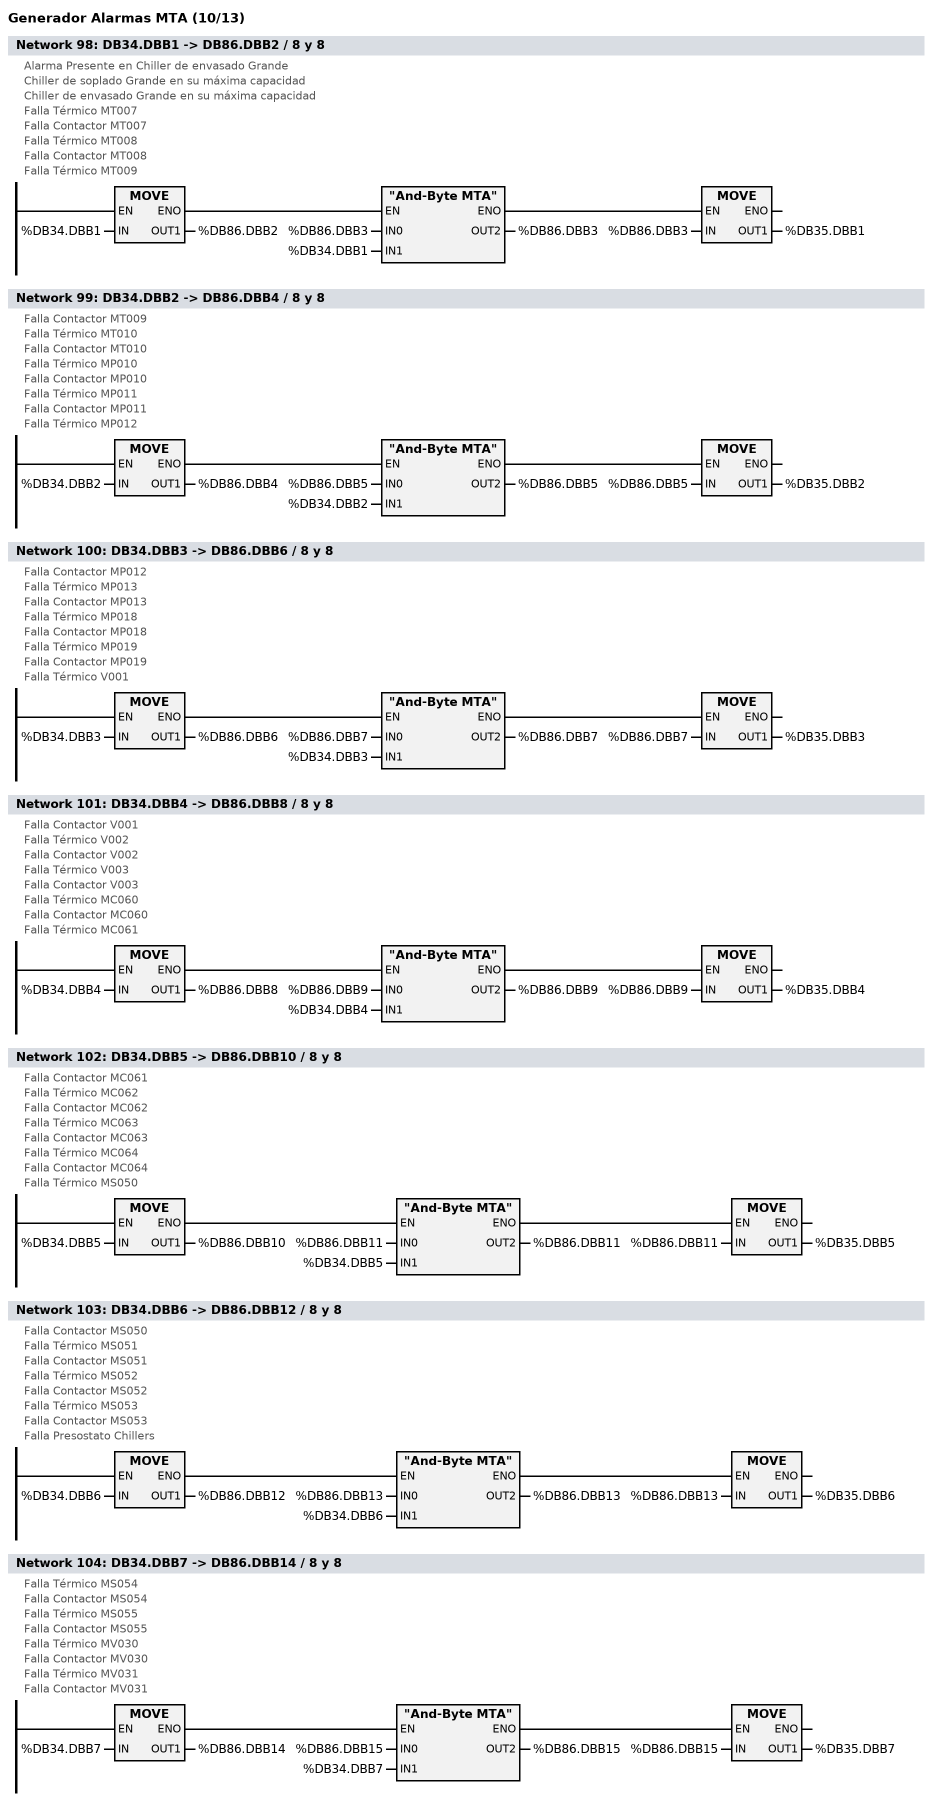
   RUNG wire#powerrail
      { S7_GenerateENO := "TRUE" } Move(in := %DB34.DBB1, out1 => %DB86.DBB2)
      "And-Byte MTA"(IN0 := %DB86.DBB3, IN1 := %DB34.DBB1, OUT2 => %DB86.DBB3)
      { S7_GenerateENO := "TRUE" } Move(in := %DB86.DBB3, out1 => %DB35.DBB1)
   END_RUNG
   // the same network as SCL:
   // ENO of a box is taken as its EN; it also drops when the box reports an error
   %DB86.DBB2 := %DB34.DBB1;
   "And-Byte MTA"(IN0 := %DB86.DBB3, IN1 := %DB34.DBB1, OUT2 => %DB86.DBB3, ENO => #_w1);
   IF #_w1 THEN %DB35.DBB1 := %DB86.DBB3; END_IF;
END_REGION

REGION Network 99: DB34.DBB2 -> DB86.DBB4 / 8 y 8
   // Falla Contactor MT009
   // Falla Térmico MT010
   // Falla Contactor MT010
   // Falla Térmico MP010
   // Falla Contactor MP010
   // Falla Térmico MP011
   // Falla Contactor MP011
   // Falla Térmico MP012
   RUNG wire#powerrail
      { S7_GenerateENO := "TRUE" } Move(in := %DB34.DBB2, out1 => %DB86.DBB4)
      "And-Byte MTA"(IN0 := %DB86.DBB5, IN1 := %DB34.DBB2, OUT2 => %DB86.DBB5)
      { S7_GenerateENO := "TRUE" } Move(in := %DB86.DBB5, out1 => %DB35.DBB2)
   END_RUNG
   // the same network as SCL:
   // ENO of a box is taken as its EN; it also drops when the box reports an error
   %DB86.DBB4 := %DB34.DBB2;
   "And-Byte MTA"(IN0 := %DB86.DBB5, IN1 := %DB34.DBB2, OUT2 => %DB86.DBB5, ENO => #_w1);
   IF #_w1 THEN %DB35.DBB2 := %DB86.DBB5; END_IF;
END_REGION

REGION Network 100: DB34.DBB3 -> DB86.DBB6 / 8 y 8
   // Falla Contactor MP012
   // Falla Térmico MP013
   // Falla Contactor MP013
   // Falla Térmico MP018
   // Falla Contactor MP018
   // Falla Térmico MP019
   // Falla Contactor MP019
   // Falla Térmico V001
   RUNG wire#powerrail
      { S7_GenerateENO := "TRUE" } Move(in := %DB34.DBB3, out1 => %DB86.DBB6)
      "And-Byte MTA"(IN0 := %DB86.DBB7, IN1 := %DB34.DBB3, OUT2 => %DB86.DBB7)
      { S7_GenerateENO := "TRUE" } Move(in := %DB86.DBB7, out1 => %DB35.DBB3)
   END_RUNG
   // the same network as SCL:
   // ENO of a box is taken as its EN; it also drops when the box reports an error
   %DB86.DBB6 := %DB34.DBB3;
   "And-Byte MTA"(IN0 := %DB86.DBB7, IN1 := %DB34.DBB3, OUT2 => %DB86.DBB7, ENO => #_w1);
   IF #_w1 THEN %DB35.DBB3 := %DB86.DBB7; END_IF;
END_REGION

REGION Network 101: DB34.DBB4 -> DB86.DBB8 / 8 y 8
   // Falla Contactor V001
   // Falla Térmico V002
   // Falla Contactor V002
   // Falla Térmico V003
   // Falla Contactor V003
   // Falla Térmico MC060
   // Falla Contactor MC060
   // Falla Térmico MC061
   RUNG wire#powerrail
      { S7_GenerateENO := "TRUE" } Move(in := %DB34.DBB4, out1 => %DB86.DBB8)
      "And-Byte MTA"(IN0 := %DB86.DBB9, IN1 := %DB34.DBB4, OUT2 => %DB86.DBB9)
      { S7_GenerateENO := "TRUE" } Move(in := %DB86.DBB9, out1 => %DB35.DBB4)
   END_RUNG
   // the same network as SCL:
   // ENO of a box is taken as its EN; it also drops when the box reports an error
   %DB86.DBB8 := %DB34.DBB4;
   "And-Byte MTA"(IN0 := %DB86.DBB9, IN1 := %DB34.DBB4, OUT2 => %DB86.DBB9, ENO => #_w1);
   IF #_w1 THEN %DB35.DBB4 := %DB86.DBB9; END_IF;
END_REGION

REGION Network 102: DB34.DBB5 -> DB86.DBB10 / 8 y 8
   // Falla Contactor MC061
   // Falla Térmico MC062
   // Falla Contactor MC062
   // Falla Térmico MC063
   // Falla Contactor MC063
   // Falla Térmico MC064
   // Falla Contactor MC064
   // Falla Térmico MS050
   RUNG wire#powerrail
      { S7_GenerateENO := "TRUE" } Move(in := %DB34.DBB5, out1 => %DB86.DBB10)
      "And-Byte MTA"(IN0 := %DB86.DBB11, IN1 := %DB34.DBB5, OUT2 => %DB86.DBB11)
      { S7_GenerateENO := "TRUE" } Move(in := %DB86.DBB11, out1 => %DB35.DBB5)
   END_RUNG
   // the same network as SCL:
   // ENO of a box is taken as its EN; it also drops when the box reports an error
   %DB86.DBB10 := %DB34.DBB5;
   "And-Byte MTA"(IN0 := %DB86.DBB11, IN1 := %DB34.DBB5, OUT2 => %DB86.DBB11, ENO => #_w1);
   IF #_w1 THEN %DB35.DBB5 := %DB86.DBB11; END_IF;
END_REGION

REGION Network 103: DB34.DBB6 -> DB86.DBB12 / 8 y 8
   // Falla Contactor MS050
   // Falla Térmico MS051
   // Falla Contactor MS051
   // Falla Térmico MS052
   // Falla Contactor MS052
   // Falla Térmico MS053
   // Falla Contactor MS053
   // Falla Presostato Chillers
   RUNG wire#powerrail
      { S7_GenerateENO := "TRUE" } Move(in := %DB34.DBB6, out1 => %DB86.DBB12)
      "And-Byte MTA"(IN0 := %DB86.DBB13, IN1 := %DB34.DBB6, OUT2 => %DB86.DBB13)
      { S7_GenerateENO := "TRUE" } Move(in := %DB86.DBB13, out1 => %DB35.DBB6)
   END_RUNG
   // the same network as SCL:
   // ENO of a box is taken as its EN; it also drops when the box reports an error
   %DB86.DBB12 := %DB34.DBB6;
   "And-Byte MTA"(IN0 := %DB86.DBB13, IN1 := %DB34.DBB6, OUT2 => %DB86.DBB13, ENO => #_w1);
   IF #_w1 THEN %DB35.DBB6 := %DB86.DBB13; END_IF;
END_REGION

REGION Network 104: DB34.DBB7 -> DB86.DBB14 / 8 y 8
   // Falla Térmico MS054
   // Falla Contactor MS054
   // Falla Térmico MS055
   // Falla Contactor MS055
   // Falla Térmico MV030
   // Falla Contactor MV030
   // Falla Térmico MV031
   // Falla Contactor MV031
   RUNG wire#powerrail
      { S7_GenerateENO := "TRUE" } Move(in := %DB34.DBB7, out1 => %DB86.DBB14)
      "And-Byte MTA"(IN0 := %DB86.DBB15, IN1 := %DB34.DBB7, OUT2 => %DB86.DBB15)
      { S7_GenerateENO := "TRUE" } Move(in := %DB86.DBB15, out1 => %DB35.DBB7)
   END_RUNG
   // the same network as SCL:
   // ENO of a box is taken as its EN; it also drops when the box reports an error
   %DB86.DBB14 := %DB34.DBB7;
   "And-Byte MTA"(IN0 := %DB86.DBB15, IN1 := %DB34.DBB7, OUT2 => %DB86.DBB15, ENO => #_w1);
   IF #_w1 THEN %DB35.DBB7 := %DB86.DBB15; END_IF;
END_REGION

REGION Network 105: DB34.DBB8 -> DB86.DBB16 / 8 y 8
   // Falla Térmico MP014
   // Falla Contactor MP014
   // Falla Térmico MP015
   // Falla Contactor MP015
   // Falla Térmico MC001
   // Falla Contactor MC001
   // Falla Térmico MC002
   // Falla Contactor MC002
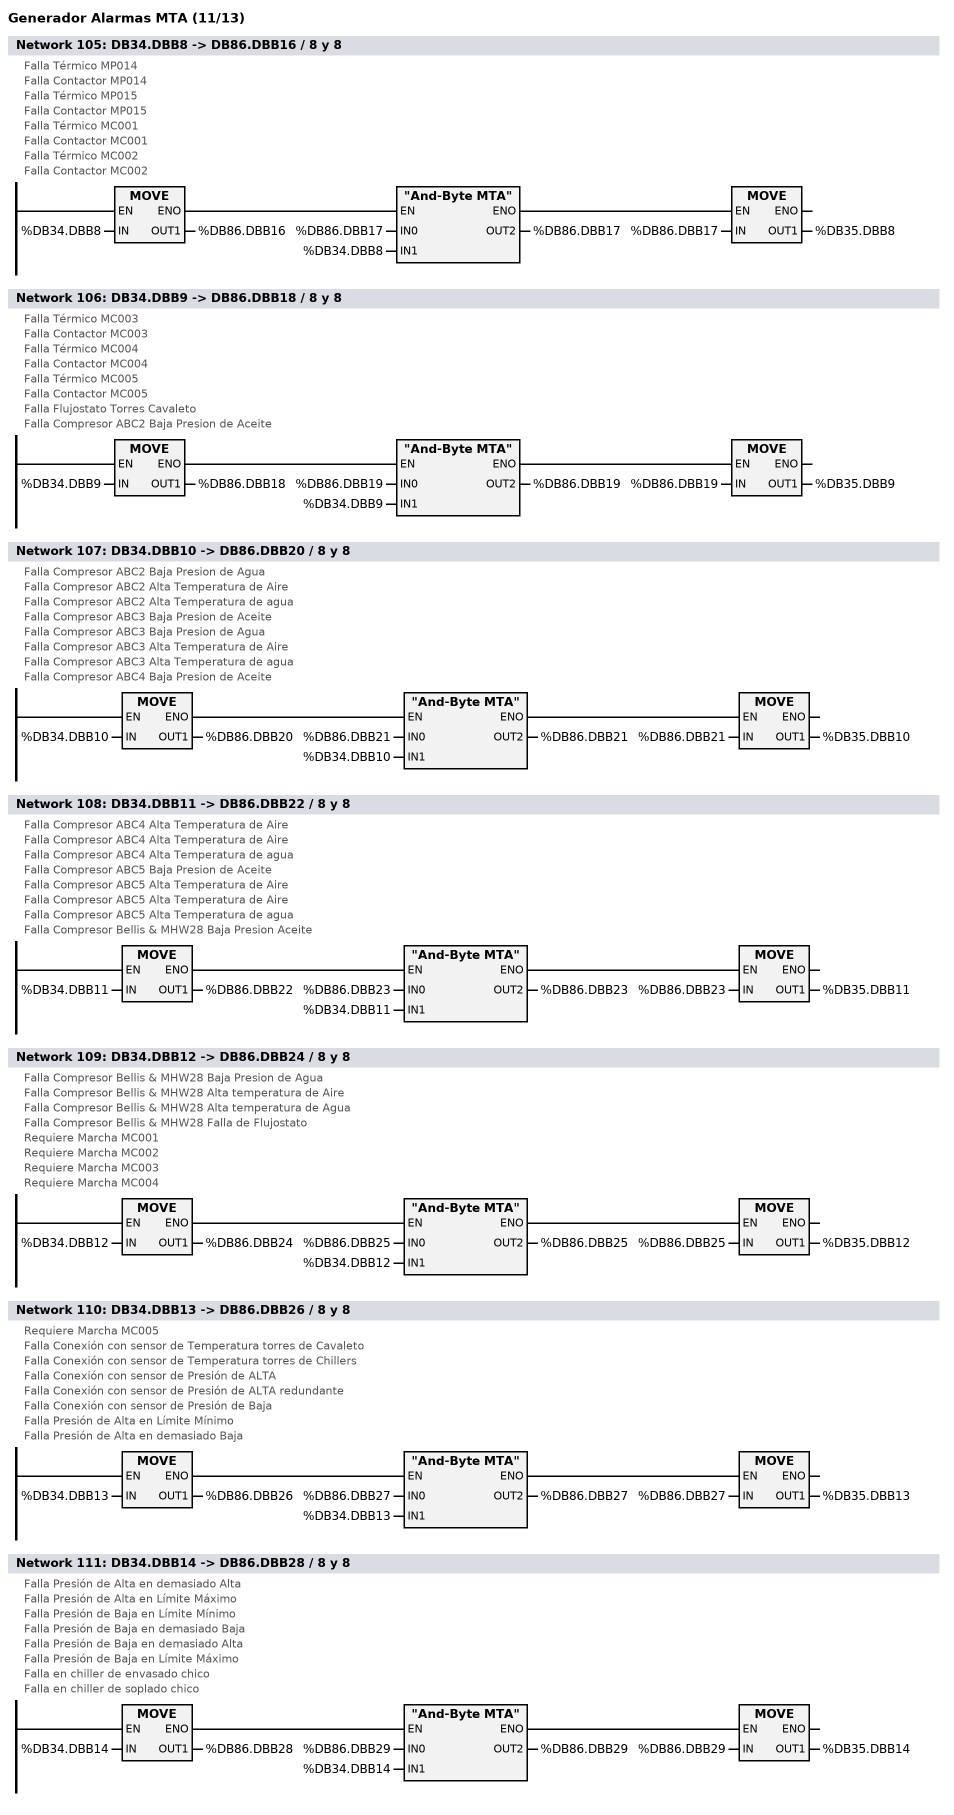
   RUNG wire#powerrail
      { S7_GenerateENO := "TRUE" } Move(in := %DB34.DBB8, out1 => %DB86.DBB16)
      "And-Byte MTA"(IN0 := %DB86.DBB17, IN1 := %DB34.DBB8, OUT2 => %DB86.DBB17)
      { S7_GenerateENO := "TRUE" } Move(in := %DB86.DBB17, out1 => %DB35.DBB8)
   END_RUNG
   // the same network as SCL:
   // ENO of a box is taken as its EN; it also drops when the box reports an error
   %DB86.DBB16 := %DB34.DBB8;
   "And-Byte MTA"(IN0 := %DB86.DBB17, IN1 := %DB34.DBB8, OUT2 => %DB86.DBB17, ENO => #_w1);
   IF #_w1 THEN %DB35.DBB8 := %DB86.DBB17; END_IF;
END_REGION

REGION Network 106: DB34.DBB9 -> DB86.DBB18 / 8 y 8
   // Falla Térmico MC003
   // Falla Contactor MC003
   // Falla Térmico MC004
   // Falla Contactor MC004
   // Falla Térmico MC005
   // Falla Contactor MC005
   // Falla Flujostato Torres Cavaleto
   // Falla Compresor ABC2 Baja Presion de Aceite
   RUNG wire#powerrail
      { S7_GenerateENO := "TRUE" } Move(in := %DB34.DBB9, out1 => %DB86.DBB18)
      "And-Byte MTA"(IN0 := %DB86.DBB19, IN1 := %DB34.DBB9, OUT2 => %DB86.DBB19)
      { S7_GenerateENO := "TRUE" } Move(in := %DB86.DBB19, out1 => %DB35.DBB9)
   END_RUNG
   // the same network as SCL:
   // ENO of a box is taken as its EN; it also drops when the box reports an error
   %DB86.DBB18 := %DB34.DBB9;
   "And-Byte MTA"(IN0 := %DB86.DBB19, IN1 := %DB34.DBB9, OUT2 => %DB86.DBB19, ENO => #_w1);
   IF #_w1 THEN %DB35.DBB9 := %DB86.DBB19; END_IF;
END_REGION

REGION Network 107: DB34.DBB10 -> DB86.DBB20 / 8 y 8
   // Falla Compresor ABC2 Baja Presion de Agua
   // Falla Compresor ABC2 Alta Temperatura de Aire
   // Falla Compresor ABC2 Alta Temperatura de agua
   // Falla Compresor ABC3 Baja Presion de Aceite
   // Falla Compresor ABC3 Baja Presion de Agua
   // Falla Compresor ABC3 Alta Temperatura de Aire
   // Falla Compresor ABC3 Alta Temperatura de agua
   // Falla Compresor ABC4 Baja Presion de Aceite
   RUNG wire#powerrail
      { S7_GenerateENO := "TRUE" } Move(in := %DB34.DBB10, out1 => %DB86.DBB20)
      "And-Byte MTA"(IN0 := %DB86.DBB21, IN1 := %DB34.DBB10, OUT2 => %DB86.DBB21)
      { S7_GenerateENO := "TRUE" } Move(in := %DB86.DBB21, out1 => %DB35.DBB10)
   END_RUNG
   // the same network as SCL:
   // ENO of a box is taken as its EN; it also drops when the box reports an error
   %DB86.DBB20 := %DB34.DBB10;
   "And-Byte MTA"(IN0 := %DB86.DBB21, IN1 := %DB34.DBB10, OUT2 => %DB86.DBB21, ENO => #_w1);
   IF #_w1 THEN %DB35.DBB10 := %DB86.DBB21; END_IF;
END_REGION

REGION Network 108: DB34.DBB11 -> DB86.DBB22 / 8 y 8
   // Falla Compresor ABC4 Alta Temperatura de Aire
   // Falla Compresor ABC4 Alta Temperatura de Aire
   // Falla Compresor ABC4 Alta Temperatura de agua
   // Falla Compresor ABC5 Baja Presion de Aceite
   // Falla Compresor ABC5 Alta Temperatura de Aire
   // Falla Compresor ABC5 Alta Temperatura de Aire
   // Falla Compresor ABC5 Alta Temperatura de agua
   // Falla Compresor Bellis & MHW28 Baja Presion Aceite
   RUNG wire#powerrail
      { S7_GenerateENO := "TRUE" } Move(in := %DB34.DBB11, out1 => %DB86.DBB22)
      "And-Byte MTA"(IN0 := %DB86.DBB23, IN1 := %DB34.DBB11, OUT2 => %DB86.DBB23)
      { S7_GenerateENO := "TRUE" } Move(in := %DB86.DBB23, out1 => %DB35.DBB11)
   END_RUNG
   // the same network as SCL:
   // ENO of a box is taken as its EN; it also drops when the box reports an error
   %DB86.DBB22 := %DB34.DBB11;
   "And-Byte MTA"(IN0 := %DB86.DBB23, IN1 := %DB34.DBB11, OUT2 => %DB86.DBB23, ENO => #_w1);
   IF #_w1 THEN %DB35.DBB11 := %DB86.DBB23; END_IF;
END_REGION

REGION Network 109: DB34.DBB12 -> DB86.DBB24 / 8 y 8
   // Falla Compresor Bellis & MHW28 Baja Presion de Agua
   // Falla Compresor Bellis & MHW28 Alta temperatura de Aire
   // Falla Compresor Bellis & MHW28 Alta temperatura de Agua
   // Falla Compresor Bellis & MHW28 Falla de Flujostato
   // Requiere Marcha MC001
   // Requiere Marcha MC002
   // Requiere Marcha MC003
   // Requiere Marcha MC004
   RUNG wire#powerrail
      { S7_GenerateENO := "TRUE" } Move(in := %DB34.DBB12, out1 => %DB86.DBB24)
      "And-Byte MTA"(IN0 := %DB86.DBB25, IN1 := %DB34.DBB12, OUT2 => %DB86.DBB25)
      { S7_GenerateENO := "TRUE" } Move(in := %DB86.DBB25, out1 => %DB35.DBB12)
   END_RUNG
   // the same network as SCL:
   // ENO of a box is taken as its EN; it also drops when the box reports an error
   %DB86.DBB24 := %DB34.DBB12;
   "And-Byte MTA"(IN0 := %DB86.DBB25, IN1 := %DB34.DBB12, OUT2 => %DB86.DBB25, ENO => #_w1);
   IF #_w1 THEN %DB35.DBB12 := %DB86.DBB25; END_IF;
END_REGION

REGION Network 110: DB34.DBB13 -> DB86.DBB26 / 8 y 8
   // Requiere Marcha MC005
   // Falla Conexión con sensor de Temperatura torres de Cavaleto
   // Falla Conexión con sensor de Temperatura torres de Chillers
   // Falla Conexión con sensor de Presión de ALTA
   // Falla Conexión con sensor de Presión de ALTA redundante
   // Falla Conexión con sensor de Presión de Baja
   // Falla Presión de Alta en Límite Mínimo
   // Falla Presión de Alta en demasiado Baja
   RUNG wire#powerrail
      { S7_GenerateENO := "TRUE" } Move(in := %DB34.DBB13, out1 => %DB86.DBB26)
      "And-Byte MTA"(IN0 := %DB86.DBB27, IN1 := %DB34.DBB13, OUT2 => %DB86.DBB27)
      { S7_GenerateENO := "TRUE" } Move(in := %DB86.DBB27, out1 => %DB35.DBB13)
   END_RUNG
   // the same network as SCL:
   // ENO of a box is taken as its EN; it also drops when the box reports an error
   %DB86.DBB26 := %DB34.DBB13;
   "And-Byte MTA"(IN0 := %DB86.DBB27, IN1 := %DB34.DBB13, OUT2 => %DB86.DBB27, ENO => #_w1);
   IF #_w1 THEN %DB35.DBB13 := %DB86.DBB27; END_IF;
END_REGION

REGION Network 111: DB34.DBB14 -> DB86.DBB28 / 8 y 8
   // Falla Presión de Alta en demasiado Alta
   // Falla Presión de Alta en Límite Máximo
   // Falla Presión de Baja en Límite Mínimo
   // Falla Presión de Baja en demasiado Baja
   // Falla Presión de Baja en demasiado Alta
   // Falla Presión de Baja en Límite Máximo
   // Falla en chiller de envasado chico
   // Falla en chiller de soplado chico
   RUNG wire#powerrail
      { S7_GenerateENO := "TRUE" } Move(in := %DB34.DBB14, out1 => %DB86.DBB28)
      "And-Byte MTA"(IN0 := %DB86.DBB29, IN1 := %DB34.DBB14, OUT2 => %DB86.DBB29)
      { S7_GenerateENO := "TRUE" } Move(in := %DB86.DBB29, out1 => %DB35.DBB14)
   END_RUNG
   // the same network as SCL:
   // ENO of a box is taken as its EN; it also drops when the box reports an error
   %DB86.DBB28 := %DB34.DBB14;
   "And-Byte MTA"(IN0 := %DB86.DBB29, IN1 := %DB34.DBB14, OUT2 => %DB86.DBB29, ENO => #_w1);
   IF #_w1 THEN %DB35.DBB14 := %DB86.DBB29; END_IF;
END_REGION

REGION Network 112: DB34.DBB15 -> DB86.DBB30 / 8 y 8
   // Horas máximas en Compresor 1
   // Horas máximas en Compresor 2
   // Horas máximas en Compresor 3
   // Horas máximas en Compresor 4
   // Horas máximas en Compresor 5
   // Falla algún contactor en Booster 1
   // Falla algún guardamotor en Booster 1
   // Presión Alta en Booster
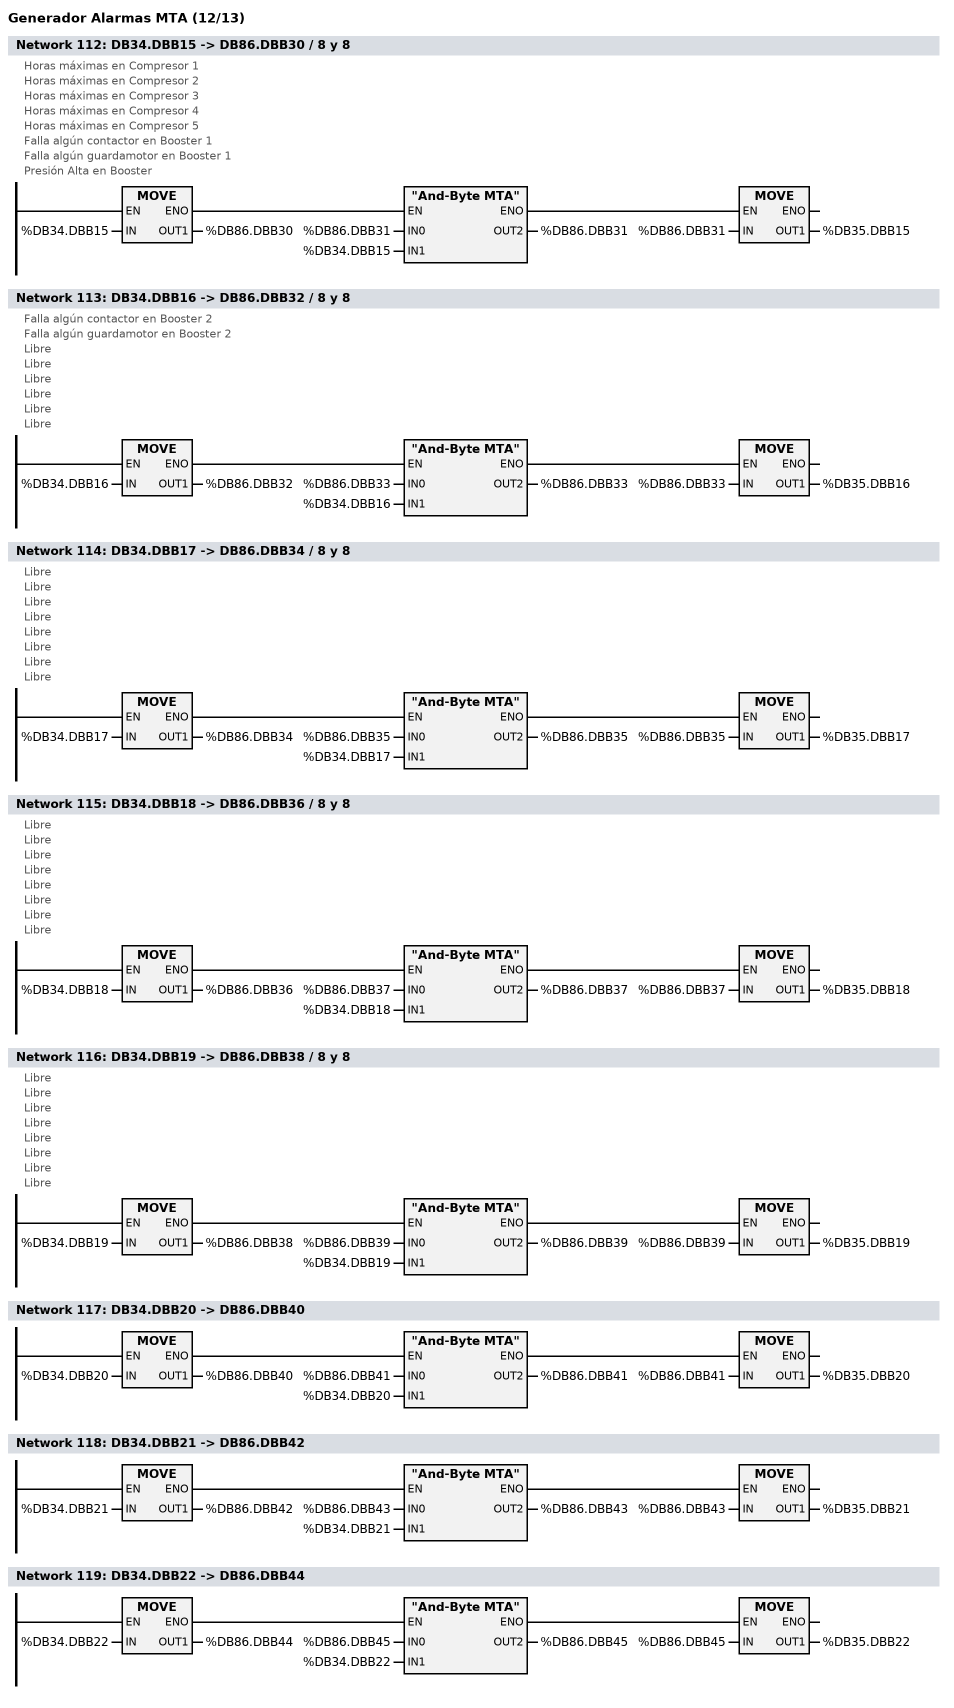
   RUNG wire#powerrail
      { S7_GenerateENO := "TRUE" } Move(in := %DB34.DBB15, out1 => %DB86.DBB30)
      "And-Byte MTA"(IN0 := %DB86.DBB31, IN1 := %DB34.DBB15, OUT2 => %DB86.DBB31)
      { S7_GenerateENO := "TRUE" } Move(in := %DB86.DBB31, out1 => %DB35.DBB15)
   END_RUNG
   // the same network as SCL:
   // ENO of a box is taken as its EN; it also drops when the box reports an error
   %DB86.DBB30 := %DB34.DBB15;
   "And-Byte MTA"(IN0 := %DB86.DBB31, IN1 := %DB34.DBB15, OUT2 => %DB86.DBB31, ENO => #_w1);
   IF #_w1 THEN %DB35.DBB15 := %DB86.DBB31; END_IF;
END_REGION

REGION Network 113: DB34.DBB16 -> DB86.DBB32 / 8 y 8
   // Falla algún contactor en Booster 2
   // Falla algún guardamotor en Booster 2
   // Libre
   // Libre
   // Libre
   // Libre
   // Libre
   // Libre
   RUNG wire#powerrail
      { S7_GenerateENO := "TRUE" } Move(in := %DB34.DBB16, out1 => %DB86.DBB32)
      "And-Byte MTA"(IN0 := %DB86.DBB33, IN1 := %DB34.DBB16, OUT2 => %DB86.DBB33)
      { S7_GenerateENO := "TRUE" } Move(in := %DB86.DBB33, out1 => %DB35.DBB16)
   END_RUNG
   // the same network as SCL:
   // ENO of a box is taken as its EN; it also drops when the box reports an error
   %DB86.DBB32 := %DB34.DBB16;
   "And-Byte MTA"(IN0 := %DB86.DBB33, IN1 := %DB34.DBB16, OUT2 => %DB86.DBB33, ENO => #_w1);
   IF #_w1 THEN %DB35.DBB16 := %DB86.DBB33; END_IF;
END_REGION

REGION Network 114: DB34.DBB17 -> DB86.DBB34 / 8 y 8
   // Libre
   // Libre
   // Libre
   // Libre
   // Libre
   // Libre
   // Libre
   // Libre
   RUNG wire#powerrail
      { S7_GenerateENO := "TRUE" } Move(in := %DB34.DBB17, out1 => %DB86.DBB34)
      "And-Byte MTA"(IN0 := %DB86.DBB35, IN1 := %DB34.DBB17, OUT2 => %DB86.DBB35)
      { S7_GenerateENO := "TRUE" } Move(in := %DB86.DBB35, out1 => %DB35.DBB17)
   END_RUNG
   // the same network as SCL:
   // ENO of a box is taken as its EN; it also drops when the box reports an error
   %DB86.DBB34 := %DB34.DBB17;
   "And-Byte MTA"(IN0 := %DB86.DBB35, IN1 := %DB34.DBB17, OUT2 => %DB86.DBB35, ENO => #_w1);
   IF #_w1 THEN %DB35.DBB17 := %DB86.DBB35; END_IF;
END_REGION

REGION Network 115: DB34.DBB18 -> DB86.DBB36 / 8 y 8
   // Libre
   // Libre
   // Libre
   // Libre
   // Libre
   // Libre
   // Libre
   // Libre
   RUNG wire#powerrail
      { S7_GenerateENO := "TRUE" } Move(in := %DB34.DBB18, out1 => %DB86.DBB36)
      "And-Byte MTA"(IN0 := %DB86.DBB37, IN1 := %DB34.DBB18, OUT2 => %DB86.DBB37)
      { S7_GenerateENO := "TRUE" } Move(in := %DB86.DBB37, out1 => %DB35.DBB18)
   END_RUNG
   // the same network as SCL:
   // ENO of a box is taken as its EN; it also drops when the box reports an error
   %DB86.DBB36 := %DB34.DBB18;
   "And-Byte MTA"(IN0 := %DB86.DBB37, IN1 := %DB34.DBB18, OUT2 => %DB86.DBB37, ENO => #_w1);
   IF #_w1 THEN %DB35.DBB18 := %DB86.DBB37; END_IF;
END_REGION

REGION Network 116: DB34.DBB19 -> DB86.DBB38 / 8 y 8
   // Libre
   // Libre
   // Libre
   // Libre
   // Libre
   // Libre
   // Libre
   // Libre
   RUNG wire#powerrail
      { S7_GenerateENO := "TRUE" } Move(in := %DB34.DBB19, out1 => %DB86.DBB38)
      "And-Byte MTA"(IN0 := %DB86.DBB39, IN1 := %DB34.DBB19, OUT2 => %DB86.DBB39)
      { S7_GenerateENO := "TRUE" } Move(in := %DB86.DBB39, out1 => %DB35.DBB19)
   END_RUNG
   // the same network as SCL:
   // ENO of a box is taken as its EN; it also drops when the box reports an error
   %DB86.DBB38 := %DB34.DBB19;
   "And-Byte MTA"(IN0 := %DB86.DBB39, IN1 := %DB34.DBB19, OUT2 => %DB86.DBB39, ENO => #_w1);
   IF #_w1 THEN %DB35.DBB19 := %DB86.DBB39; END_IF;
END_REGION

REGION Network 117: DB34.DBB20 -> DB86.DBB40
   RUNG wire#powerrail
      { S7_GenerateENO := "TRUE" } Move(in := %DB34.DBB20, out1 => %DB86.DBB40)
      "And-Byte MTA"(IN0 := %DB86.DBB41, IN1 := %DB34.DBB20, OUT2 => %DB86.DBB41)
      { S7_GenerateENO := "TRUE" } Move(in := %DB86.DBB41, out1 => %DB35.DBB20)
   END_RUNG
   // the same network as SCL:
   // ENO of a box is taken as its EN; it also drops when the box reports an error
   %DB86.DBB40 := %DB34.DBB20;
   "And-Byte MTA"(IN0 := %DB86.DBB41, IN1 := %DB34.DBB20, OUT2 => %DB86.DBB41, ENO => #_w1);
   IF #_w1 THEN %DB35.DBB20 := %DB86.DBB41; END_IF;
END_REGION

REGION Network 118: DB34.DBB21 -> DB86.DBB42
   RUNG wire#powerrail
      { S7_GenerateENO := "TRUE" } Move(in := %DB34.DBB21, out1 => %DB86.DBB42)
      "And-Byte MTA"(IN0 := %DB86.DBB43, IN1 := %DB34.DBB21, OUT2 => %DB86.DBB43)
      { S7_GenerateENO := "TRUE" } Move(in := %DB86.DBB43, out1 => %DB35.DBB21)
   END_RUNG
   // the same network as SCL:
   // ENO of a box is taken as its EN; it also drops when the box reports an error
   %DB86.DBB42 := %DB34.DBB21;
   "And-Byte MTA"(IN0 := %DB86.DBB43, IN1 := %DB34.DBB21, OUT2 => %DB86.DBB43, ENO => #_w1);
   IF #_w1 THEN %DB35.DBB21 := %DB86.DBB43; END_IF;
END_REGION

REGION Network 119: DB34.DBB22 -> DB86.DBB44
   RUNG wire#powerrail
      { S7_GenerateENO := "TRUE" } Move(in := %DB34.DBB22, out1 => %DB86.DBB44)
      "And-Byte MTA"(IN0 := %DB86.DBB45, IN1 := %DB34.DBB22, OUT2 => %DB86.DBB45)
      { S7_GenerateENO := "TRUE" } Move(in := %DB86.DBB45, out1 => %DB35.DBB22)
   END_RUNG
   // the same network as SCL:
   // ENO of a box is taken as its EN; it also drops when the box reports an error
   %DB86.DBB44 := %DB34.DBB22;
   "And-Byte MTA"(IN0 := %DB86.DBB45, IN1 := %DB34.DBB22, OUT2 => %DB86.DBB45, ENO => #_w1);
   IF #_w1 THEN %DB35.DBB22 := %DB86.DBB45; END_IF;
END_REGION

REGION Network 120: DB34.DBB23 -> DB86.DBB46
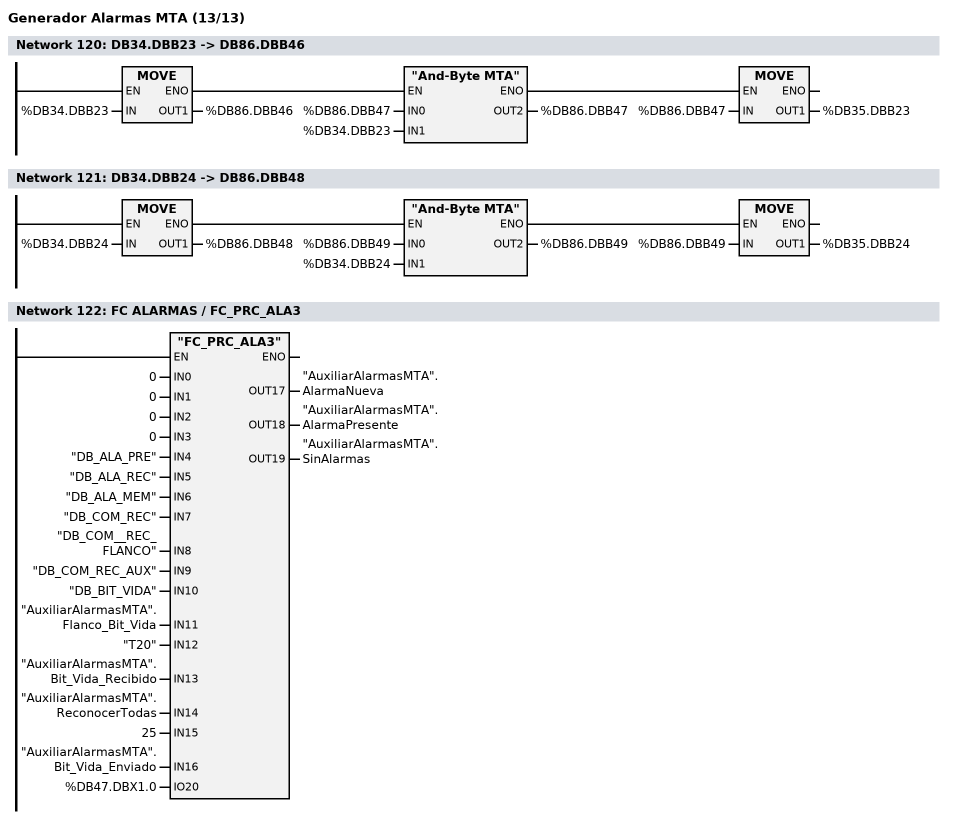
   RUNG wire#powerrail
      { S7_GenerateENO := "TRUE" } Move(in := %DB34.DBB23, out1 => %DB86.DBB46)
      "And-Byte MTA"(IN0 := %DB86.DBB47, IN1 := %DB34.DBB23, OUT2 => %DB86.DBB47)
      { S7_GenerateENO := "TRUE" } Move(in := %DB86.DBB47, out1 => %DB35.DBB23)
   END_RUNG
   // the same network as SCL:
   // ENO of a box is taken as its EN; it also drops when the box reports an error
   %DB86.DBB46 := %DB34.DBB23;
   "And-Byte MTA"(IN0 := %DB86.DBB47, IN1 := %DB34.DBB23, OUT2 => %DB86.DBB47, ENO => #_w1);
   IF #_w1 THEN %DB35.DBB23 := %DB86.DBB47; END_IF;
END_REGION

REGION Network 121: DB34.DBB24 -> DB86.DBB48
   RUNG wire#powerrail
      { S7_GenerateENO := "TRUE" } Move(in := %DB34.DBB24, out1 => %DB86.DBB48)
      "And-Byte MTA"(IN0 := %DB86.DBB49, IN1 := %DB34.DBB24, OUT2 => %DB86.DBB49)
      { S7_GenerateENO := "TRUE" } Move(in := %DB86.DBB49, out1 => %DB35.DBB24)
   END_RUNG
   // the same network as SCL:
   // ENO of a box is taken as its EN; it also drops when the box reports an error
   %DB86.DBB48 := %DB34.DBB24;
   "And-Byte MTA"(IN0 := %DB86.DBB49, IN1 := %DB34.DBB24, OUT2 => %DB86.DBB49, ENO => #_w1);
   IF #_w1 THEN %DB35.DBB24 := %DB86.DBB49; END_IF;
END_REGION

REGION Network 122: FC ALARMAS / FC_PRC_ALA3
   RUNG wire#powerrail
      "FC_PRC_ALA3"(IN0 := 0, IN1 := 0, IN2 := 0, IN3 := 0, IN4 := "DB_ALA_PRE", IN5 := "DB_ALA_REC", IN6 := "DB_ALA_MEM", IN7 := "DB_COM_REC", IN8 := "DB_COM__REC_FLANCO", IN9 := "DB_COM_REC_AUX", IN10 := "DB_BIT_VIDA", IN11 := "AuxiliarAlarmasMTA".Flanco_Bit_Vida, IN12 := "T20", IN13 := "AuxiliarAlarmasMTA".Bit_Vida_Recibido, IN14 := "AuxiliarAlarmasMTA".ReconocerTodas, IN15 := 25, IN16 := "AuxiliarAlarmasMTA".Bit_Vida_Enviado, IO20 := %DB47.DBX1.0, OUT17 => "AuxiliarAlarmasMTA".AlarmaNueva, OUT18 => "AuxiliarAlarmasMTA".AlarmaPresente, OUT19 => "AuxiliarAlarmasMTA".SinAlarmas)
   END_RUNG
   // the same network as SCL:
   "FC_PRC_ALA3"(IN0 := 0,
                 IN1 := 0,
                 IN2 := 0,
                 IN3 := 0,
                 IN4 := "DB_ALA_PRE",
                 IN5 := "DB_ALA_REC",
                 IN6 := "DB_ALA_MEM",
                 IN7 := "DB_COM_REC",
                 IN8 := "DB_COM__REC_FLANCO",
                 IN9 := "DB_COM_REC_AUX",
                 IN10 := "DB_BIT_VIDA",
                 IN11 := "AuxiliarAlarmasMTA".Flanco_Bit_Vida,
                 IN12 := "T20",
                 IN13 := "AuxiliarAlarmasMTA".Bit_Vida_Recibido,
                 IN14 := "AuxiliarAlarmasMTA".ReconocerTodas,
                 IN15 := 25,
                 IN16 := "AuxiliarAlarmasMTA".Bit_Vida_Enviado,
                 IO20 := %DB47.DBX1.0,
                 OUT17 => "AuxiliarAlarmasMTA".AlarmaNueva,
                 OUT18 => "AuxiliarAlarmasMTA".AlarmaPresente,
                 OUT19 => "AuxiliarAlarmasMTA".SinAlarmas);
END_REGION
END_FUNCTION

FUNCTION "FalCmpAlta" : Void   // FC49, LAD
{ S7_Optimized_Access := 'FALSE' }
VERSION : 0.1
   VAR_TEMP   // added for the SCL form of the ladder/FBD networks
      _w1 : Bool;
      _w2 : Bool;
      _s5time1 : S5Time;
   END_VAR
BEGIN

REGION Network 1: Fallas de MC001 - Compresor de Alta ABC2
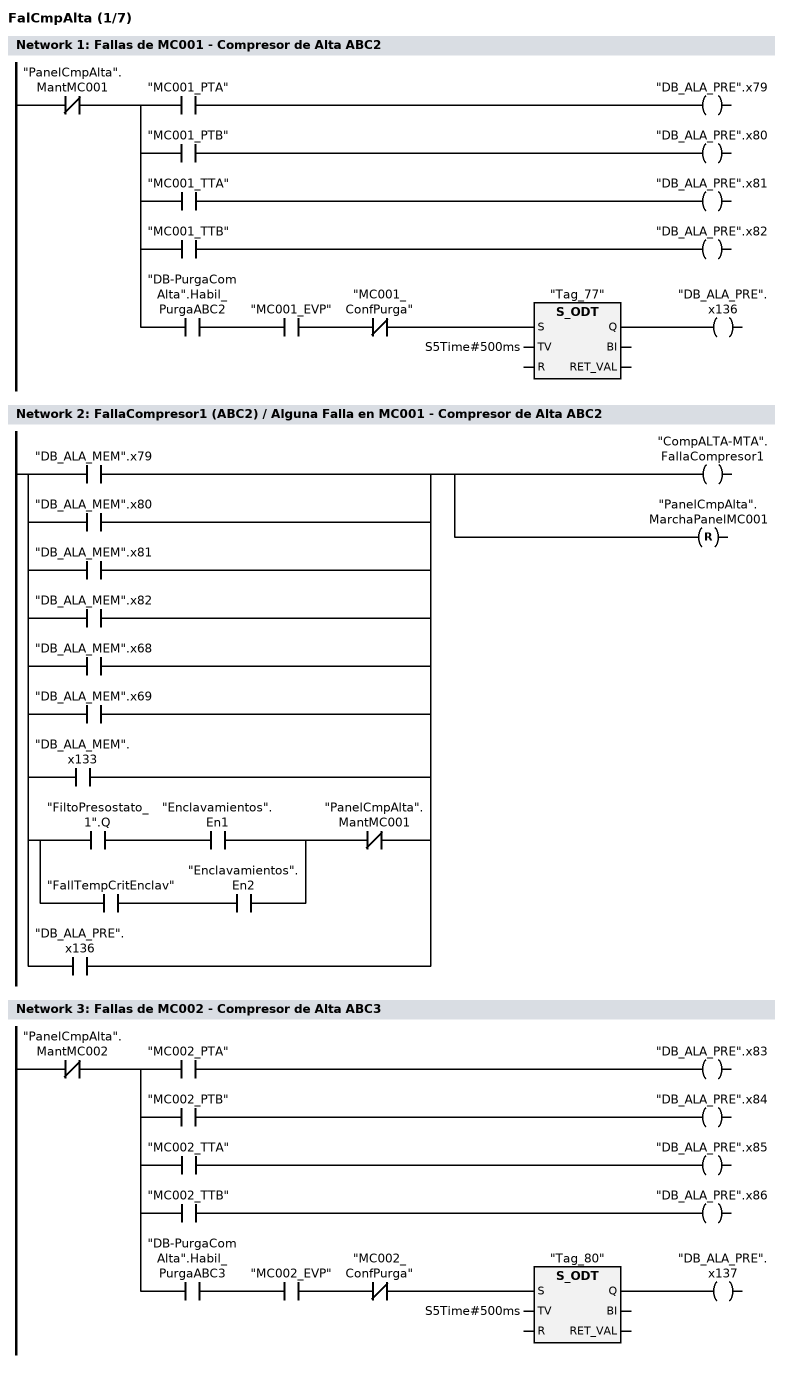
   RUNG wire#powerrail
      I_Contact( "PanelCmpAlta".MantMC001 )
      wire#w1
      Contact( "MC001_PTA" )
      Coil( "DB_ALA_PRE".x79 )
   END_RUNG
   RUNG wire#w1
      Contact( "MC001_PTB" )
      Coil( "DB_ALA_PRE".x80 )
   END_RUNG
   RUNG wire#w1
      Contact( "MC001_TTA" )
      Coil( "DB_ALA_PRE".x81 )
   END_RUNG
   RUNG wire#w1
      Contact( "MC001_TTB" )
      Coil( "DB_ALA_PRE".x82 )
   END_RUNG
   RUNG wire#w1
      Contact( "DB-PurgaComAlta".Habil_PurgaABC2 )
      Contact( "MC001_EVP" )
      I_Contact( "MC001_ConfPurga" )
      S_ODT(T_NO := "Tag_77", TV := S5Time#500ms, R :=, BI =>, RET_VAL =>)
      Coil( "DB_ALA_PRE".x136 )
   END_RUNG
   // the same network as SCL:
   #_w1 := NOT "PanelCmpAlta".MantMC001;
   "DB_ALA_PRE".x79 := #_w1 AND "MC001_PTA";
   "DB_ALA_PRE".x80 := #_w1 AND "MC001_PTB";
   "DB_ALA_PRE".x81 := #_w1 AND "MC001_TTA";
   "DB_ALA_PRE".x82 := #_w1 AND "MC001_TTB";
   #_s5time1 := S_ODT(T_NO := "Tag_77",
                      S := #_w1 AND "DB-PurgaComAlta".Habil_PurgaABC2 AND "MC001_EVP" AND NOT "MC001_ConfPurga",
                      TV := S5Time#500ms,
                      Q => #_w2);
   "DB_ALA_PRE".x136 := #_w2;
END_REGION

REGION Network 2: FallaCompresor1 (ABC2) / Alguna Falla en MC001 - Compresor de Alta ABC2
   RUNG wire#powerrail
      Contact( "DB_ALA_MEM".x79 )
      wire#w1
      Coil( "CompALTA-MTA".FallaCompresor1 )
   END_RUNG
   RUNG wire#powerrail
      Contact( "DB_ALA_MEM".x80 )
   END_RUNG wire#w1
   RUNG wire#powerrail
      Contact( "DB_ALA_MEM".x81 )
   END_RUNG wire#w1
   RUNG wire#powerrail
      Contact( "DB_ALA_MEM".x82 )
   END_RUNG wire#w1
   RUNG wire#powerrail
      Contact( "DB_ALA_MEM".x68 )
   END_RUNG wire#w1
   RUNG wire#powerrail
      Contact( "DB_ALA_MEM".x69 )
   END_RUNG wire#w1
   RUNG wire#powerrail
      Contact( "DB_ALA_MEM".x133 )
   END_RUNG wire#w1
   RUNG wire#powerrail
      Contact( "FiltoPresostato_1".Q )
      Contact( "Enclavamientos".En1 )
      wire#w2
      I_Contact( "PanelCmpAlta".MantMC001 )
   END_RUNG wire#w1
   RUNG wire#powerrail
      Contact( "FallTempCritEnclav" )
      Contact( "Enclavamientos".En2 )
   END_RUNG wire#w2
   RUNG wire#powerrail
      Contact( "DB_ALA_PRE".x136 )
   END_RUNG wire#w1
   RUNG wire#w1
      R_Coil( "PanelCmpAlta".MarchaPanelMC001 )
   END_RUNG
   // the same network as SCL:
   "CompALTA-MTA".FallaCompresor1 := "DB_ALA_MEM".x79 OR "DB_ALA_MEM".x80 OR "DB_ALA_MEM".x81 OR "DB_ALA_MEM".x82 OR "DB_ALA_MEM".x68 OR "DB_ALA_MEM".x69 OR "DB_ALA_MEM".x133 OR ((("FiltoPresostato_1".Q AND "Enclavamientos".En1) OR ("FallTempCritEnclav" AND "Enclavamientos".En2)) AND NOT "PanelCmpAlta".MantMC001) OR "DB_ALA_PRE".x136;
   IF "CompALTA-MTA".FallaCompresor1 THEN "PanelCmpAlta".MarchaPanelMC001 := FALSE; END_IF;
END_REGION

REGION Network 3: Fallas de MC002 - Compresor de Alta ABC3
   RUNG wire#powerrail
      I_Contact( "PanelCmpAlta".MantMC002 )
      wire#w1
      Contact( "MC002_PTA" )
      Coil( "DB_ALA_PRE".x83 )
   END_RUNG
   RUNG wire#w1
      Contact( "MC002_PTB" )
      Coil( "DB_ALA_PRE".x84 )
   END_RUNG
   RUNG wire#w1
      Contact( "MC002_TTA" )
      Coil( "DB_ALA_PRE".x85 )
   END_RUNG
   RUNG wire#w1
      Contact( "MC002_TTB" )
      Coil( "DB_ALA_PRE".x86 )
   END_RUNG
   RUNG wire#w1
      Contact( "DB-PurgaComAlta".Habil_PurgaABC3 )
      Contact( "MC002_EVP" )
      I_Contact( "MC002_ConfPurga" )
      S_ODT(T_NO := "Tag_80", TV := S5Time#500ms, R :=, BI =>, RET_VAL =>)
      Coil( "DB_ALA_PRE".x137 )
   END_RUNG
   // the same network as SCL:
   #_w1 := NOT "PanelCmpAlta".MantMC002;
   "DB_ALA_PRE".x83 := #_w1 AND "MC002_PTA";
   "DB_ALA_PRE".x84 := #_w1 AND "MC002_PTB";
   "DB_ALA_PRE".x85 := #_w1 AND "MC002_TTA";
   "DB_ALA_PRE".x86 := #_w1 AND "MC002_TTB";
   #_s5time1 := S_ODT(T_NO := "Tag_80",
                      S := #_w1 AND "DB-PurgaComAlta".Habil_PurgaABC3 AND "MC002_EVP" AND NOT "MC002_ConfPurga",
                      TV := S5Time#500ms,
                      Q => #_w2);
   "DB_ALA_PRE".x137 := #_w2;
END_REGION

REGION Network 4: FallaCompresor2 (ABC3) / Alguna Falla en MC002 - Compresor de Alta ABC3